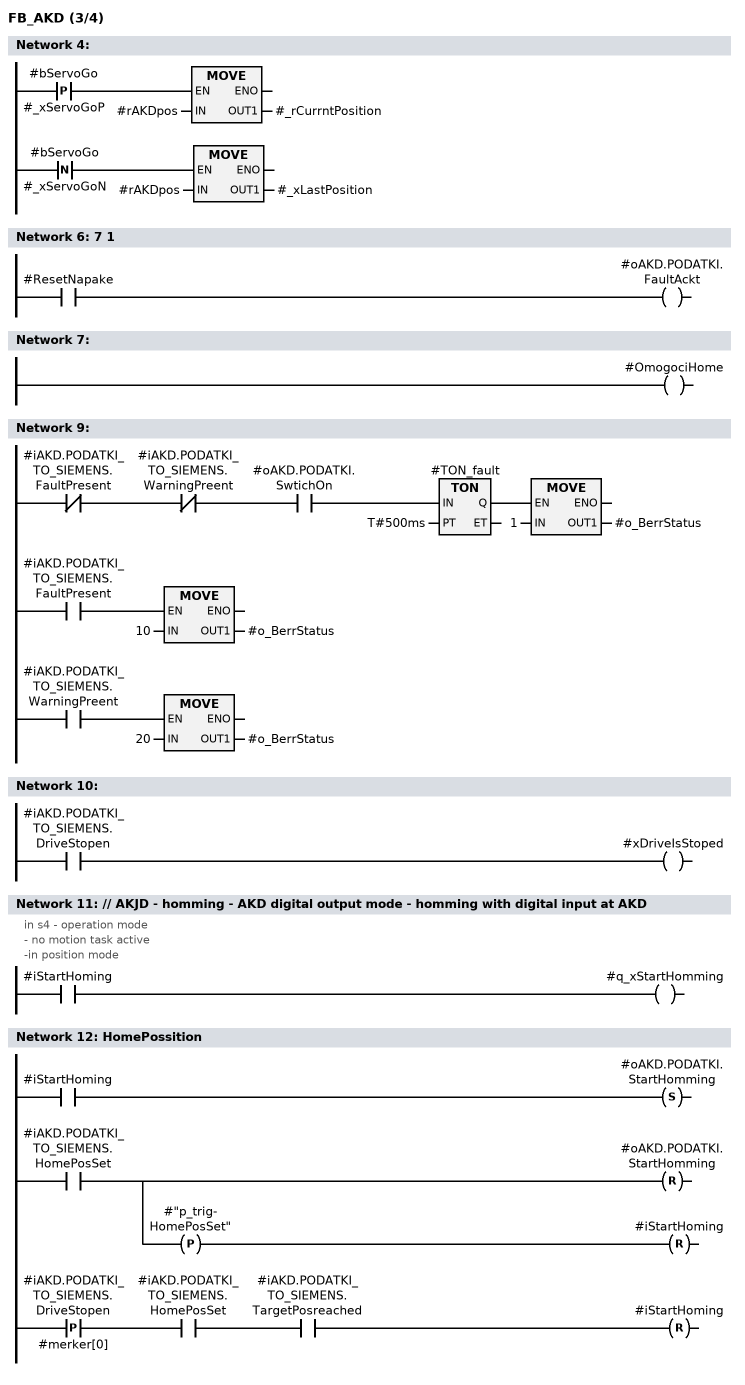
   RUNG wire#powerrail
      P_Contact(operand := #bServoGo, bit := #_xServoGoP)
      Move(in := #rAKDpos, out1 => #_rCurrntPosition)
   END_RUNG
   RUNG wire#powerrail
      N_Contact(operand := #bServoGo, bit := #_xServoGoN)
      Move(in := #rAKDpos, out1 => #_xLastPosition)
   END_RUNG
   // the same network as SCL:
   #_w1 := #bServoGo AND NOT #_xServoGoP;   // rising edge of #bServoGo
   #_xServoGoP := #bServoGo;
   IF #_w1 THEN #_rCurrntPosition := #rAKDpos; END_IF;
   #_w2 := NOT #bServoGo AND #_xServoGoN;   // falling edge of #bServoGo
   #_xServoGoN := #bServoGo;
   IF #_w2 THEN #_xLastPosition := #rAKDpos; END_IF;
END_REGION

REGION Network 5 (SCL)
   //PretvorbaHitrosti
   #diHitrost := INT_TO_REAL(#iNastavitevHitrosti);
   #dwHitrostRez :=((#diHitrost * 4294967295/12000));
   #oAKD.PODATKI.MDI_VELOCITY := REAL_TO_DINT(#dwHitrostRez); //hitrost


   // Operation mode
   #oAKD.PODATKI.MDI_MOD := 16#00_00; //0 - relativni 1//aboslutni gib
   #oAKD.PODATKI.SATANW := #iStPrograma;   //OutputTask

   //pretvorba poziij
   #AKDcurrPos := (#iAKD.PODATKI_TO_SIEMENS.ActualPos * 5 )/ 65536;
   #rAKDpos:= (#iAKD.PODATKI_TO_SIEMENS.ActualPos) / 65536.00;
   //nastavljanjePozicije
   //nastavljanje pozicije
   #oAKD.PODATKI.MDI_TARPOS := (65536 * #dNastavitevPozicije / 5);
END_REGION

REGION Network 6: 7 1
   RUNG wire#powerrail
      Contact( #ResetNapake )
      Coil( #oAKD.PODATKI.FaultAckt )
   END_RUNG
   // the same network as SCL:
   #oAKD.PODATKI.FaultAckt := #ResetNapake;
END_REGION

REGION Network 7
   RUNG wire#powerrail
      Coil( #OmogociHome )
   END_RUNG
   // the same network as SCL:
   #OmogociHome := TRUE;
END_REGION

REGION Network 8: ERROR STATUS
END_REGION

REGION Network 9
   #TON_fault(IN := NOT #iAKD.PODATKI_TO_SIEMENS.FaultPresent AND NOT #iAKD.PODATKI_TO_SIEMENS.WarningPreent AND #oAKD.PODATKI.SwtichOn,   // TON
              PT := T#500ms);
   IF #TON_fault.Q THEN #o_BerrStatus := 1; END_IF;
   IF #iAKD.PODATKI_TO_SIEMENS.FaultPresent THEN #o_BerrStatus := 10; END_IF;
   IF #iAKD.PODATKI_TO_SIEMENS.WarningPreent THEN #o_BerrStatus := 20; END_IF;
END_REGION

REGION Network 10
   RUNG wire#powerrail
      Contact( #iAKD.PODATKI_TO_SIEMENS.DriveStopen )
      Coil( #xDriveIsStoped )
   END_RUNG
   // the same network as SCL:
   #xDriveIsStoped := #iAKD.PODATKI_TO_SIEMENS.DriveStopen;
END_REGION

REGION Network 11: // AKJD - homming - AKD digital output mode - homming with digital input at AKD
   // in s4 - operation mode
   // - no motion task active
   // -in position mode
   RUNG wire#powerrail
      Contact( #iStartHoming )
      Coil( #q_xStartHomming )
   END_RUNG
   // the same network as SCL:
   #q_xStartHomming := #iStartHoming;
END_REGION

REGION Network 12: HomePossition
   RUNG wire#powerrail
      Contact( #iStartHoming )
      S_Coil( #oAKD.PODATKI.StartHomming )
   END_RUNG
   RUNG wire#powerrail
      Contact( #iAKD.PODATKI_TO_SIEMENS.HomePosSet )
      wire#w1
      R_Coil( #oAKD.PODATKI.StartHomming )
   END_RUNG
   RUNG wire#w1
      P_Trig( #"p_trig-HomePosSet" )
      R_Coil( #iStartHoming )
   END_RUNG
   RUNG wire#powerrail
      P_Contact(operand := #iAKD.PODATKI_TO_SIEMENS.DriveStopen, bit := #merker[0])
      Contact( #iAKD.PODATKI_TO_SIEMENS.HomePosSet )
      Contact( #iAKD.PODATKI_TO_SIEMENS.TargetPosreached )
      R_Coil( #iStartHoming )
   END_RUNG
   // the same network as SCL:
   IF #iStartHoming THEN #oAKD.PODATKI.StartHomming := TRUE; END_IF;
   IF #iAKD.PODATKI_TO_SIEMENS.HomePosSet THEN #oAKD.PODATKI.StartHomming := FALSE; END_IF;
   #_w1 := #iAKD.PODATKI_TO_SIEMENS.HomePosSet AND NOT #"p_trig-HomePosSet";   // rising edge
   #"p_trig-HomePosSet" := #iAKD.PODATKI_TO_SIEMENS.HomePosSet;
   IF #_w1 THEN #iStartHoming := FALSE; END_IF;
   #_w2 := #iAKD.PODATKI_TO_SIEMENS.DriveStopen AND NOT #merker[0];   // rising edge of #iAKD.PODATKI_TO_SIEMENS.DriveStopen
   #merker[0] := #iAKD.PODATKI_TO_SIEMENS.DriveStopen;
   IF #_w2 AND #iAKD.PODATKI_TO_SIEMENS.HomePosSet AND #iAKD.PODATKI_TO_SIEMENS.TargetPosreached THEN
       #iStartHoming := FALSE;
   END_IF;
END_REGION

REGION Network 13: OUTPUT : is hommed
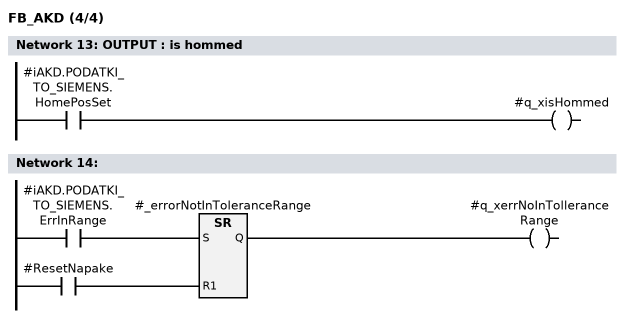
   RUNG wire#powerrail
      Contact( #iAKD.PODATKI_TO_SIEMENS.HomePosSet )
      Coil( #q_xisHommed )
   END_RUNG
   // the same network as SCL:
   #q_xisHommed := #iAKD.PODATKI_TO_SIEMENS.HomePosSet;
END_REGION

REGION Network 14
   RUNG wire#powerrail
      Contact( #iAKD.PODATKI_TO_SIEMENS.ErrInRange )
      S_SR(operand := #_errorNotInToleranceRange, r1 := wire#w1)
      Coil( #q_xerrNoInTolleranceRange )
   END_RUNG
   RUNG wire#powerrail
      Contact( #ResetNapake )
   END_RUNG wire#w1
   // the same network as SCL:
   IF #iAKD.PODATKI_TO_SIEMENS.ErrInRange THEN
       #_errorNotInToleranceRange := TRUE;   // SR flip-flop
   END_IF;
   IF #ResetNapake THEN #_errorNotInToleranceRange := FALSE; END_IF;
   #q_xerrNoInTolleranceRange := #_errorNotInToleranceRange;
END_REGION
END_FUNCTION_BLOCK

FUNCTION_BLOCK "AKD_PN_TG400_v05"   // FB14, SCL
TITLE = AKD_PN_TG400_TIA13_v05
{ S7_Optimized_Access := 'FALSE' }
AUTHOR : jcoleman
FAMILY : TG400
VERSION : 5.0
// This function block supports Profinet communication with the AKD drive using Telegram 400.  It is written in TIA V13. 
// For more information, please see the AKD Profinet Manual and the supporting documentation for this function block.
   VAR_INPUT
      iID : Hw_Io;   // Hardware identifier
      iInit : Bool;   // initialize config for TG400
      iEStop : Bool;   // immediate quick stop and disable
      iSW_Enable : Bool;   // enable/disable
      iStop : Bool;   // stop all movement
      iReset : Bool;   // reset drive faults
      iStart_Homing : Bool;   // start homing
      iStart_Jog : Bool;   // start jog
      iStart_Move : Bool;   // start motion task
      iMT_Pause : Bool;   // pause active motion task
      iMT_MoveType : Word;   // motion task control word 0 = relative; 1 = absolute
      iMTNum : Word;   // motion task number 0x8000 = direct motion task
      iCmdPos : DWord;   // commanded position for motion task or homing
      iCmdVel : DWord;   // commanded velocity for jog or direct motion task
      iCmdAcc : Word;   // commanded acceleration for jog or direct motion task
      iCmdDec : Word;   // commanded deceleration for jog or direct motion task
   END_VAR
   VAR_OUTPUT
      oInitDone : Bool;   // initialization status - 0 while configuring TG400, 1= done
      oStatus : DWord;   // ZSW1
      oPos : DWord;   // actual position
      oVel : Word;   // actual velocity x * 12000 rpm / 2^15
      oCurrent : Word;   // actual current x *DRV.IPEAK / 2^14
      oEnabled : Bool;   // Drive power on
      oError : Bool;   // fault in function block or communication
      oMoving : Bool;   // axis enabled and moving
      oHomed : Bool;   // axis homed
      oInPos : Bool;   // axis within in-position window
      oFault : Bool;   // drive fault
      oWarning : Bool;   // drive warning
   END_VAR
   VAR
      TG_400 : "UDT_AKD_TG400";
      wPNReadStatus : Word;
      bPNReadError : Bool;
      wPNWriteStatus : Word;
      bPNWriteError : Bool;
      bResetDone : Bool;
      bHomeStarted : Bool;
      bStartMoveDone : Bool;
      bEstop : Bool;
      wStartReset : Int;
      wStartMove : Int;
      wSDOStatus : Word;
      bySDODataArray : Array[0..63] of Byte;
      SDOWrite : WRREC;
      SDORead : RDREC;
      bSDOReq : Bool;
      bSDOWriteBusy : Bool;
      bSDOWriteDone : Bool;
      bSDOWriteError : Bool;
      bSDOReadBusy : Bool;
      bSDOReadDone : Bool;
      bSDOReadError : Bool;
      wSDOReadValue : Word;
      wSDOAddress : Word;
      bSWEnabled : Bool;
      wHomingStartPoint : Word;
      bStartMove : Bool;
      bSDOStatusReadActive : Bool;
   END_VAR
BEGIN
   ////////////////////////////////////////////////////////////////////////////////////////////////////////
   // Standard communication module between a Kollmorgen AKD and S7-1200/1500 PLC
   //
   // Version  When        Who         What
   // ---------------------------------------------
   // V 05     09.05.17    JColeman KM Changed Telegram 400 mapping PNU writes to be individual writes, rather
   //                                  than a block write...to be more robust.
   // V 04     08.31.17    JColeman KM Changed error handling to indicate internal block errors.
   // V 03     06.05.17    JColeman KM Changed EStop code to set flag without waiting for motion to stop. 
   //                                  Added setting opmode=2 in init section.
   //                                  Added comments.
   //                                  Added information to FB properties.
   //                                  Turn on real-time jog mode during enable process.
   //                                  Do not use Optimized block access.
   // V 02     05.12.17    JColeman KM Changed names of inputs and outputs to be more user friendly
   //                                  Added output oInitDone to indicate when the telegram configuration is complete
   //                                  Changed name of FB to be specific to TG400
   //                                  Changed verion numbering
   // V 1.000  17.09.15    MRupf KM    Conversion to TIA V13 SP1
   // V 0.004  09.07.15    MRupf KM    Home_dist changed to DINT variable length
   //          06.07.15    MRupf KM    Fault and Warning read locked angainst interruption
   // V 0.003  05.06.15    MRupf KM    New iStart_MT is only accepted after the ZSW1 Bit 12 is FALSE again
   //          03.06.15    MRupf KM    Handshake to start motion task with ZSW1 Bit 12 and auto reset after 500ms #285
   //          14.04.15    MRupf KM    Init write cases extended to not do endless recall on error
   //                                  Homing start stop bug, #246-250
   //                                  Reset STW1.6/.7 only after two PN cylce #214, 283
   // V 0.002  26.02.15    MRupf KM    Setup Telegramm 400 with HOME.DIST, VL.FB, IL.FB
   //                                  Read Fault and Warning No. if acitve
   //                                  Reset STW if drive fault happens while enabled    
   // V 0.001  18.02.15    MRupf KM    First version
   //////////////////////////////////////////////////////////////////////////////////////////////////////////

   // initialisation
   IF #iInit THEN
       #wSDOStatus := 0;
       #oInitDone := FALSE;    //False during telegram configuration
   END_IF;
   IF #wSDOStatus < 20 THEN //set telegram send data = 0
       #TG_400.Send.STW1 := 0;
       #TG_400.Send.SATZANW := 0;
       #TG_400.Send.STW2 := 0;
       #TG_400.Send.MDI_TARPOS := 0;
       #TG_400.Send.MDI_VELOCITY := 0;
       #TG_400.Send.MDI_ACC := 0;
       #TG_400.Send.MDI_DEC := 0;
       #TG_400.Send.MDI_MOD := 0;

       #bPNReadError := FALSE;
       #bPNWriteError := FALSE;
   END_IF;

   // Do the setup of the Telegram 400
   IF NOT #iInit AND #wSDOStatus < 19 THEN

       // Map Telegram 400 Send
       // Clear the Array and start the request
       IF #wSDOStatus = 0 THEN
           FILL_BLK(IN := 0,
                    COUNT := 64,
                    OUT => #bySDODataArray[0]);
           #bSDOReq := TRUE;
           #bSDOWriteDone := FALSE;
           #wSDOStatus := 1; //proceed to Step 1
       END_IF;
       // setup the array data and start WRREC
       IF #wSDOStatus = 1 THEN //Step 1
           #bySDODataArray[0] := 16#ff; //Request Reference
           #bySDODataArray[1] := 16#02; //2 for write PNU
           #bySDODataArray[2] := 16#00; //Axis# is 0 for AKD
           #bySDODataArray[3] := 16#01; //number of parameters
           // Set PNU 915 subindex 8
           #bySDODataArray[4] := 16#10; //Attribute is 0x10
           #bySDODataArray[5] := 16#01; //Number of elements =1
           #bySDODataArray[6] := 16#03; //0x393 for PNU 915
           #bySDODataArray[7] := 16#93; //PNU 915
           #bySDODataArray[8] := 16#00; //subindex
           #bySDODataArray[9] := 16#08; //subindex 8 for 8th word of telegram
           // To PNU 100 (HOME.DIST)
           #bySDODataArray[10] := 16#42; //Format =0x42 for Word
           #bySDODataArray[11] := 16#01; //Number of values
           #bySDODataArray[12] := 16#00; //data
           #bySDODataArray[13] := 16#64; //data - Signal #100 for HOME.DIST

           #SDOWrite(REQ := #bSDOReq, //do the PNU write
                     ID := #iID,
                     INDEX := 47, //AKD suppors "Record Data 47"
                     LEN := 14,   //data length
                     BUSY => #bSDOWriteBusy,
                     DONE => #bSDOWriteDone,
                     ERROR => #bSDOWriteError,
                     RECORD := #bySDODataArray);
           IF #bSDOWriteBusy THEN
               #bSDOReq := FALSE;
           ELSIF #bSDOWriteDone THEN
               #wSDOStatus := 2; //proceed to Step 2
           END_IF;
       END_IF;

       // Map Telegram 400 Receive
       // Clear the Array and start the request
       IF #wSDOStatus = 2 THEN //Step 2
           FILL_BLK(IN := 0,
                    COUNT := 64,
                    OUT => #bySDODataArray[0]);
           #bSDOReq := TRUE;
           #bSDOWriteDone := FALSE;
           #wSDOStatus := 3; //proceed to Step 3
       END_IF;
       // setup the array data and start WRREC
       IF #wSDOStatus = 3 THEN //Step 3
           #bySDODataArray[0] := 16#fe; //Request Reference
           #bySDODataArray[1] := 16#02; //2 for write PNU
           #bySDODataArray[2] := 16#00; //Axis# is 0 for AKD
           #bySDODataArray[3] := 16#01; // Number of parameters to write at a time
           // Set PNU 916 subindex 0
           #bySDODataArray[4] := 16#10; //Attribute is 0x10
           #bySDODataArray[5] := 16#01; //Number of elements =1
           #bySDODataArray[6] := 16#03; //0x394 for PNU 916
           #bySDODataArray[7] := 16#94; //PNU 916
           #bySDODataArray[8] := 16#00; //subindex
           #bySDODataArray[9] := 16#00; //subindex 0 for 1st word of telegram
           // To PNU 2 (ZSW1)
           #bySDODataArray[10] := 16#42; //Format =0x42 for Word
           #bySDODataArray[11] := 16#01; //Number of values
           #bySDODataArray[12] := 16#00; //data
           #bySDODataArray[13] := 16#02; //data - Signal #2 (0x02) for ZSW1

           #SDOWrite(REQ := #bSDOReq, //do the PNU write
                     ID := #iID,
                     INDEX := 47, //AKD suppors "Record Data 47"
                     LEN := 14,   //data length
                     BUSY => #bSDOWriteBusy,
                     DONE => #bSDOWriteDone,
                     ERROR => #bSDOWriteError,
                     RECORD := #bySDODataArray);
           IF #bSDOWriteBusy THEN
               #bSDOReq := FALSE;
           ELSIF #bSDOWriteDone THEN
               #wSDOStatus := 4; //proceed to Step 4
           END_IF;
       END_IF;

       // Clear the Array and start the request
       IF #wSDOStatus = 4 THEN //Step 4
           FILL_BLK(IN := 0,
                    COUNT := 64,
                    OUT => #bySDODataArray[0]);
           #bSDOReq := TRUE;
           #bSDOWriteDone := FALSE;
           #wSDOStatus := 5; //proceed to Step 5
       END_IF;
       // setup the array data and start WRREC
       IF #wSDOStatus = 5 THEN //Step 5
           #bySDODataArray[0] := 16#fd; //Request Reference
           #bySDODataArray[1] := 16#02; //2 for write PNU
           #bySDODataArray[2] := 16#00; //Axis# is 0 for AKD
           #bySDODataArray[3] := 16#01; // Number of parameters to write at a time
           // Set PNU 916 subindex 1
           #bySDODataArray[4] := 16#10; //Attribute is 0x10
           #bySDODataArray[5] := 16#01; //Number of elements =1
           #bySDODataArray[6] := 16#03; //0x394 for PNU 916
           #bySDODataArray[7] := 16#94; //PNU 916
           #bySDODataArray[8] := 16#00; //subindex
           #bySDODataArray[9] := 16#01; //subindex 1 for 2nd word of telegram
           // To PNU 33 (AKTSATZ)
           #bySDODataArray[10] := 16#42; //Format =0x42 for Word
           #bySDODataArray[11] := 16#01; //Number of values
           #bySDODataArray[12] := 16#00; //data
           #bySDODataArray[13] := 16#21; //data - Signal #33 (0x21) for AKTSATZ

           #SDOWrite(REQ := #bSDOReq, //do the PNU write
                     ID := #iID,
                     INDEX := 47, //AKD suppors "Record Data 47"
                     LEN := 14,   //data length
                     BUSY => #bSDOWriteBusy,
                     DONE => #bSDOWriteDone,
                     ERROR => #bSDOWriteError,
                     RECORD := #bySDODataArray);
           IF #bSDOWriteBusy THEN
               #bSDOReq := FALSE;
           ELSIF #bSDOWriteDone THEN
               #wSDOStatus := 6; //proceed to Step 6
           END_IF;
       END_IF;

       // Clear the Array and start the request
       IF #wSDOStatus = 6 THEN //Step 6
           FILL_BLK(IN := 0,
                    COUNT := 64,
                    OUT => #bySDODataArray[0]);
           #bSDOReq := TRUE;
           #bSDOWriteDone := FALSE;
           #wSDOStatus := 7; //proceed to Step 7
       END_IF;
       // setup the array data and start WRREC
       IF #wSDOStatus = 7 THEN //Step 7
           #bySDODataArray[0] := 16#fc; //Request Reference
           #bySDODataArray[1] := 16#02; //2 for write PNU
           #bySDODataArray[2] := 16#00; //Axis# is 0 for AKD
           #bySDODataArray[3] := 16#01; // Number of parameters to write at a time
           // Set PNU 916 subindex 2
           #bySDODataArray[4] := 16#10; //Attribute is 0x10
           #bySDODataArray[5] := 16#01; //Number of elements =1
           #bySDODataArray[6] := 16#03; //0x394 for PNU 916
           #bySDODataArray[7] := 16#94; //PNU 916
           #bySDODataArray[8] := 16#00; //subindex
           #bySDODataArray[9] := 16#02; //subindex 2 for 3rd word of telegram
           // To PNU 4 (ZSW1)
           #bySDODataArray[10] := 16#42; //Format =0x42 for Word
           #bySDODataArray[11] := 16#01; //Number of values
           #bySDODataArray[12] := 16#00; //data
           #bySDODataArray[13] := 16#04; //data - Signal #4 (0x04) for ZSW2

           #SDOWrite(REQ := #bSDOReq, //do the PNU write
                     ID := #iID,
                     INDEX := 47, //AKD suppors "Record Data 47"
                     LEN := 14,   //data length
                     BUSY => #bSDOWriteBusy,
                     DONE => #bSDOWriteDone,
                     ERROR => #bSDOWriteError,
                     RECORD := #bySDODataArray);
           IF #bSDOWriteBusy THEN
               #bSDOReq := FALSE;
           ELSIF #bSDOWriteDone THEN
               #wSDOStatus := 8; //proceed to Step 8
           END_IF;
       END_IF;

       // Clear the Array and start the request
       IF #wSDOStatus = 8 THEN //Step 8
           FILL_BLK(IN := 0,
                    COUNT := 64,
                    OUT => #bySDODataArray[0]);
           #bSDOReq := TRUE;
           #bSDOWriteDone := FALSE;
           #wSDOStatus := 9; //proceed to Step 9
       END_IF;
       // setup the array data and start WRREC
       IF #wSDOStatus = 9 THEN //Step 9
           #bySDODataArray[0] := 16#fb; //Request Reference
           #bySDODataArray[1] := 16#02; //2 for write PNU
           #bySDODataArray[2] := 16#00; //Axis# is 0 for AKD
           #bySDODataArray[3] := 16#01; // Number of parameters to write at a time
           // Set PNU 916 subindex 3
           #bySDODataArray[4] := 16#10; //Attribute is 0x10
           #bySDODataArray[5] := 16#01; //Number of elements =1
           #bySDODataArray[6] := 16#03; //0x394 for PNU 916
           #bySDODataArray[7] := 16#94; //PNU 916
           #bySDODataArray[8] := 16#00; //subindex
           #bySDODataArray[9] := 16#03; //subindex 3 for 4th word of telegram
           // To PNU 28 (XIST_A)
           #bySDODataArray[10] := 16#42; //Format =0x42 for Word
           #bySDODataArray[11] := 16#01; //Number of values
           #bySDODataArray[12] := 16#00; //data
           #bySDODataArray[13] := 16#1C; //data - Signal #28 (0x1C) for XIST_A

           #SDOWrite(REQ := #bSDOReq, //do the PNU write
                     ID := #iID,
                     INDEX := 47, //AKD suppors "Record Data 47"
                     LEN := 14,   //data length
                     BUSY => #bSDOWriteBusy,
                     DONE => #bSDOWriteDone,
                     ERROR => #bSDOWriteError,
                     RECORD := #bySDODataArray);
           IF #bSDOWriteBusy THEN
               #bSDOReq := FALSE;
           ELSIF #bSDOWriteDone THEN
               #wSDOStatus := 10; //proceed to Step 10
           END_IF;
       END_IF;

       // Clear the Array and start the request
       IF #wSDOStatus = 10 THEN //Step 10
           FILL_BLK(IN := 0,
                    COUNT := 64,
                    OUT => #bySDODataArray[0]);
           #bSDOReq := TRUE;
           #bSDOWriteDone := FALSE;
           #wSDOStatus := 11; //proceed to Step 11
       END_IF;
       // setup the array data and start WRREC
       IF #wSDOStatus = 11 THEN //Step 11
           #bySDODataArray[0] := 16#fa; //Request Reference
           #bySDODataArray[1] := 16#02; //2 for write PNU
           #bySDODataArray[2] := 16#00; //Axis# is 0 for AKD
           #bySDODataArray[3] := 16#01; // Number of parameters to write at a time
           // Set PNU 916 subindex 4
           #bySDODataArray[4] := 16#10; //Attribute is 0x10
           #bySDODataArray[5] := 16#01; //Number of elements =1
           #bySDODataArray[6] := 16#03; //0x394 for PNU 916
           #bySDODataArray[7] := 16#94; //PNU 916
           #bySDODataArray[8] := 16#00; //subindex
           #bySDODataArray[9] := 16#04; //subindex 4 for 5th word of telegram
           // To PNU 6 (NIST_A)
           #bySDODataArray[10] := 16#42; //Format =0x42 for Word
           #bySDODataArray[11] := 16#01; //Number of values
           #bySDODataArray[12] := 16#00; //data
           #bySDODataArray[13] := 16#06; //data - Signal #6 (0x06) for NIST_A (VL.FB)

           #SDOWrite(REQ := #bSDOReq, //do the PNU write
                     ID := #iID,
                     INDEX := 47, //AKD suppors "Record Data 47"
                     LEN := 14,   //data length
                     BUSY => #bSDOWriteBusy,
                     DONE => #bSDOWriteDone,
                     ERROR => #bSDOWriteError,
                     RECORD := #bySDODataArray);
           IF #bSDOWriteBusy THEN
               #bSDOReq := FALSE;
           ELSIF #bSDOWriteDone THEN
               #wSDOStatus := 12; //proceed to Step 12
           END_IF;
       END_IF;

       // Clear the Array and start the request
       IF #wSDOStatus = 12 THEN //Step 12
           FILL_BLK(IN := 0,
                    COUNT := 64,
                    OUT => #bySDODataArray[0]);
           #bSDOReq := TRUE;
           #bSDOWriteDone := FALSE;
           #wSDOStatus := 13; //proceed to Step 13
       END_IF;
       // setup the array data and start WRREC
       IF #wSDOStatus = 13 THEN //Step 13
           #bySDODataArray[0] := 16#f9; //Request Reference
           #bySDODataArray[1] := 16#02; //2 for write PNU
           #bySDODataArray[2] := 16#00; //Axis# is 0 for AKD
           #bySDODataArray[3] := 16#01; // Number of parameters to write at a time
           // Set PNU 916 subindex 5
           #bySDODataArray[4] := 16#10; //Attribute is 0x10
           #bySDODataArray[5] := 16#01; //Number of elements =1
           #bySDODataArray[6] := 16#03; //0x394 for PNU 916
           #bySDODataArray[7] := 16#94; //PNU 916
           #bySDODataArray[8] := 16#00; //subindex
           #bySDODataArray[9] := 16#05; //subindex 5 for 6th word of telegram
           // To PNU 52 (ITIST_GLATT)
           #bySDODataArray[10] := 16#42; //Format =0x42 for Word
           #bySDODataArray[11] := 16#01; //Number of values
           #bySDODataArray[12] := 16#00; //data
           #bySDODataArray[13] := 16#34; //data - Signal #52 (0x34) for ITIST_GLATT (IL.FB)

           #SDOWrite(REQ := #bSDOReq, //do the PNU write
                     ID := #iID,
                     INDEX := 47, //AKD suppors "Record Data 47"
                     LEN := 14,   //data length
                     BUSY => #bSDOWriteBusy,
                     DONE => #bSDOWriteDone,
                     ERROR => #bSDOWriteError,
                     RECORD := #bySDODataArray);
           IF #bSDOWriteBusy THEN
               #bSDOReq := FALSE;
           ELSIF #bSDOWriteDone THEN
               #wSDOStatus := 14; //proceed to Step 14
               //#oInitDone := 1;    //telegram configuration complete
           END_IF;
       END_IF;

       // Set OpMode 
       // Clear the Array and start the request
       IF #wSDOStatus = 14 THEN //Step 14
           FILL_BLK(IN := 0,
                    COUNT := 64,
                    OUT => #bySDODataArray[0]);
           #bSDOReq := TRUE;
           #bSDOWriteDone := FALSE;
           #wSDOStatus := 15; //proceed to Step 15
       END_IF;
       // Set OpMode = 2 Position
       IF #wSDOStatus = 15 THEN //Step 15
           #bySDODataArray[0] := 16#fe; //Request Reference
           #bySDODataArray[1] := 16#02; //2 for write PNU
           #bySDODataArray[2] := 16#00; //Axis# is 0 for AKD
           #bySDODataArray[3] := 16#01; // Number of parameters to write at a time
               // Set PNU 930 subindex 0 (DRV.OPMODE)
           #bySDODataArray[4] := 16#10; //Attribute is 0x10
           #bySDODataArray[5] := 16#01; //Number of elements =1
           #bySDODataArray[6] := 16#03; //0x3A2 for PNU 930 - opmode
           #bySDODataArray[7] := 16#A2; //PNU 930
           #bySDODataArray[8] := 16#00; //subindex 0
           #bySDODataArray[9] := 16#00; //subindex 0
               // To 2 (position mode)
           #bySDODataArray[10] := 16#42; //Format =0x42 for Word
           #bySDODataArray[11] := 16#01; //Number of values
           #bySDODataArray[12] := 16#02; //data
           #bySDODataArray[13] := 16#02; //data - vlaue = 2 for position mode

           #SDOWrite(REQ := #bSDOReq, //do the PNU write
                     ID := #iID,
                     INDEX := 47, //AKD suppors "Record Data 47"
                     LEN := 14,   //data length
                     BUSY => #bSDOWriteBusy,
                     DONE => #bSDOWriteDone,
                     ERROR => #bSDOWriteError,
                     RECORD := #bySDODataArray);
           IF #bSDOWriteBusy THEN
               #bSDOReq := FALSE;
           ELSIF #bSDOWriteDone THEN
               #wSDOStatus := 20; // setup complete - skip to process
               #oInitDone := TRUE;    //telegram configuration complete
           END_IF;
       END_IF;
   END_IF;

   // Read ZSW and set output values
   IF NOT #iInit AND #wSDOStatus > 19 THEN
       #wPNReadStatus := DPRD_DAT(LADDR := #iID,
                                  RECORD => #TG_400.Receive);
       IF #wPNReadStatus = 0 THEN
           #bPNReadError := FALSE;

           #oStatus.%W0 := #TG_400.Receive.ZSW1;
           IF #wSDOStatus > 20 THEN
               #oStatus.%W1 := #wSDOReadValue;
           ELSE
               #oStatus.%W1 := 0;
           END_IF;
           #oPos.%W0 := #TG_400.Receive.XIST_A_1;
           #oPos.%W1 := #TG_400.Receive.XIST_A;
           #oVel := #TG_400.Receive.NIST_A;
           #oCurrent := #TG_400.Receive.ITIST_GLATT;

           #oEnabled := #TG_400.Receive.ZSW1.%X0 AND #TG_400.Receive.ZSW1.%X1 AND #TG_400.Receive.ZSW1.%X2 AND NOT #TG_400.Receive.ZSW1.%X6;
           #oFault := #TG_400.Receive.ZSW1.%X3;
           #oMoving := NOT #TG_400.Receive.ZSW1.%X13 OR #TG_400.Receive.ZSW1.%X14 OR #TG_400.Receive.ZSW1.%X12;
           #oHomed := #TG_400.Receive.ZSW1.%X11;
           IF #TG_400.Send.STW1.%X6 THEN        // Reset the InPos Flag for a minimum of one write cycle
               #oInPos := FALSE;
           ELSE
               #oInPos := #TG_400.Receive.ZSW1.%X10;
           END_IF;
           #oWarning := #TG_400.Receive.ZSW1.%X7;
       ELSE
           #bPNReadError := TRUE;
       END_IF;

   END_IF;

   // Do the write always as the zero Telegramm needs to be send on a init aswell
   #wPNWriteStatus := DPWR_DAT(LADDR := #iID,
                               RECORD := #TG_400.Send);

   // set STW1 and values for the AKD
   IF NOT #iInit AND #wSDOStatus > 19 THEN
       IF #wPNWriteStatus = 0 THEN
           #bPNWriteError := FALSE;

           #TG_400.Send.STW1.%X10 := TRUE;
           IF #TG_400.Receive.ZSW1.%X9 THEN     // PLC has control

               // Do a EStop
               IF #iEStop THEN
                   #TG_400.Send.STW1.%X2 := FALSE;
                   #bEstop := TRUE;
               END_IF;

               // Do a reset
               IF #iReset AND NOT #bResetDone THEN
                   #wSDOStatus := 20;
                   #TG_400.Send.STW1.%X7 := TRUE;
                   #bResetDone := TRUE;
                   #bEstop := FALSE;
                   #wStartReset := #TG_400.Receive.ZSW2;
               END_IF;
               IF ABS(#wStartReset - #TG_400.Receive.ZSW2) > 2 THEN
                   #TG_400.Send.STW1.%X7 := FALSE;
               END_IF;

               // Enable the drive
               IF #iSW_Enable AND NOT #bEstop AND NOT (#bSWEnabled AND #TG_400.Receive.ZSW1.%X6 OR #TG_400.Receive.ZSW1.%X3) THEN
                   IF #TG_400.Receive.ZSW1.%X6 THEN      // Switch on inhibited
                       #TG_400.Send.STW1.%X1 := TRUE;
                       #TG_400.Send.STW1.%X2 := TRUE;
                   ELSE
                       IF #TG_400.Receive.ZSW1.%X0 THEN     // Ready for switiching on
                           #TG_400.Send.STW1.%X0 := TRUE;
                           IF #TG_400.Receive.ZSW1.%X1 THEN       // Switched on
                               #TG_400.Send.STW1.%X3 := TRUE;
                               IF #TG_400.Receive.ZSW1.%X2 THEN       // Operation
                                   #TG_400.Send.STW1.%X12 := TRUE; //turn on real time jogging mode
                                   #bSWEnabled := TRUE;

                                   // Do a Stop
                                   IF #iStop THEN
                                       #TG_400.Send.STW1.%X4 := FALSE;   // Stop active motion task
                                       #TG_400.Send.STW1.%X5 := FALSE;   // Stop active motion task
                                       #TG_400.Send.STW1.%X8 := FALSE;   // Stop jog 1
                                       #TG_400.Send.STW1.%X9 := FALSE;   // Stop jog 2
                                       #TG_400.Send.STW1.%X11 := FALSE;  // Stop homeing
                                       //#TG_400.Send.STW1.%X12 := FALSE;  // Stop real time jogging mode
                                   ELSE

                                       // Do home
                                       IF #iStart_Homing AND NOT #bHomeStarted THEN
                                           #TG_400.Send.HOME_DIST := #iCmdPos.%W1;
                                           #TG_400.Send.HOME_DIST_1 := #iCmdPos.%W0;
                                           #TG_400.Send.STW1.%X11 := TRUE;
                                           #wHomingStartPoint := #TG_400.Receive.ZSW2;
                                           #bHomeStarted := TRUE;
                                       ELSE
                                           IF #TG_400.Receive.ZSW1.%X11 AND #TG_400.Receive.ZSW1.%X13 AND (ABS(#wHomingStartPoint - #TG_400.Receive.ZSW2) > 5) THEN
                                               #TG_400.Send.STW1.%X11 := FALSE;
                                           END_IF;

                                           // Jogging
                                           IF #iStart_Jog AND #iCmdVel <> 0 THEN
                                               #TG_400.Send.STW1.%X8 := TRUE;
                                               //#TG_400.Send.STW1.%X12 := TRUE;

                                               // if the speed input is negative set Bit 13 for reverse direction 
                                               IF #iCmdVel.%X31 = 1 THEN
                                                   #TG_400.Send.STW1.%X13 := TRUE;
                                                   #TG_400.Send.MDI_VELOCITY := (16#ffff - #iCmdVel.%W1 + 1);
                                                   #TG_400.Send.MDI_VELOCITY_1 := (16#ffff - #iCmdVel.%W0 + 1);
                                               ELSE
                                                   #TG_400.Send.STW1.%X13 := FALSE;
                                                   #TG_400.Send.MDI_VELOCITY := #iCmdVel.%W1;
                                                   #TG_400.Send.MDI_VELOCITY_1 := #iCmdVel.%W0;
                                               END_IF;

                                               #TG_400.Send.MDI_ACC := #iCmdAcc;
                                               #TG_400.Send.MDI_DEC := #iCmdDec;
                                           ELSE
                                               #TG_400.Send.STW1.%X8 := FALSE;
                                               //#TG_400.Send.STW1.%X12 := FALSE;

                                               // Interrupt a move
                                               IF #iMT_Pause THEN
                                                   #TG_400.Send.STW1.%X5 := FALSE;    // intermediate stop, motion is paused and will continue when the pause is lifted
                                               ELSE
                                                   #TG_400.Send.STW1.%X5 := TRUE;    // No intermediate stop
                                               END_IF;

                                               // Reset the rising edge of the start bit to be read for the next task
                                               IF #TG_400.Receive.ZSW1.%X12 OR ABS(#wStartMove - #TG_400.Receive.ZSW2) > 62 THEN //if start command has been acknowledged, or >62 telegram transmissions
                                                   #bStartMoveDone := TRUE; // the process to start the move has been completed
                                                   #TG_400.Send.STW1.%X6 := FALSE; //turn off the start bit
                                               END_IF;
                                               // Move
                                               IF #iStart_Move AND NOT #bStartMove THEN
                                                   #TG_400.Send.MDI_MOD := #iMT_MoveType;   // 1 = absolute, 0 = relative
                                                   #TG_400.Send.SATZANW := #iMTNum;      // 0x8000 = direct motion task, otherwise select a motion task from the AKD
                                                   #TG_400.Send.MDI_TARPOS := #iCmdPos.%W1;
                                                   #TG_400.Send.MDI_TARPOS_1 := #iCmdPos.%W0;
                                                   #TG_400.Send.MDI_VELOCITY := #iCmdVel.%W1;
                                                   #TG_400.Send.MDI_VELOCITY_1 := #iCmdVel.%W0;
                                                   #TG_400.Send.MDI_ACC := #iCmdAcc;
                                                   #TG_400.Send.MDI_DEC := #iCmdDec;
                                                   #TG_400.Send.STW1.%X4 := TRUE;    // Do not reject traversing task
                                                   #TG_400.Send.STW1.%X5 := TRUE;    // No intermediate stop
                                                   #TG_400.Send.STW1.%X6 := TRUE;    // Start the move

                                                   #bStartMove := TRUE; // the process to start the move has been started but not completed
                                                   #bStartMoveDone := FALSE; // the process to start the move has not been completed
                                                   #wStartMove := #TG_400.Receive.ZSW2;
                                               END_IF; //If Start move

                                           END_IF; //If Start Jog
                                       END_IF; //If Start Homing
                                   END_IF; // If Stop
                               END_IF; // If ZSW1 bit2 Operation Enabled
                           END_IF; // If ZSW1 bit1 Switched On
                       END_IF; // If ZSW1 bit0 Ready for Switch On
                   END_IF; // If ZSW1 bit6 Switch-On Inhibited

                   // If the axis gets disabled all the corresponding motion signals have to be reset    
               ELSE
                   #bSWEnabled := FALSE;

                   #TG_400.Send.STW1.%X0 := FALSE;
                   #TG_400.Send.STW1.%X1 := FALSE;
                   #TG_400.Send.STW1.%X2 := FALSE;
                   #TG_400.Send.STW1.%X3 := FALSE;
                   #TG_400.Send.STW1.%X4 := FALSE;
                   #TG_400.Send.STW1.%X5 := FALSE;
                   #TG_400.Send.STW1.%X6 := FALSE;
                   #TG_400.Send.STW1.%X8 := FALSE;
                   #TG_400.Send.STW1.%X9 := FALSE;
                   #TG_400.Send.STW1.%X11 := FALSE;
                   #TG_400.Send.STW1.%X12 := FALSE;
               END_IF; //If Enable
           END_IF; // ZSW1 bit9 PLC has control
       ELSE
           #bPNWriteError := TRUE;
       END_IF; //If #wPNWriteStatus = 0

       // Read drive faults and warning on occurens
       IF #oFault THEN
           // If alarm is not read yet: start read
           IF NOT #wSDOStatus.%X6 AND NOT #bSDOStatusReadActive THEN
               #wSDOStatus := 64;
               #wSDOAddress := 16#09AD;     // Read PNU 2477 (DRV.FAULT1)
               #bSDOStatusReadActive := TRUE;
           END_IF;

           // If warning is not read yet: start read
       ELSIF #oWarning THEN
           IF NOT #wSDOStatus.%X5 AND NOT #bSDOStatusReadActive THEN
               #wSDOStatus := 32;
               #wSDOAddress := 16#0AE7;    // Read PNU2791 (DRV.WARNING1)
               #bSDOStatusReadActive := TRUE;
           END_IF;
       ELSE
           IF NOT #bSDOStatusReadActive THEN
               #wSDOStatus := 20;
           END_IF;
       END_IF; //IF #oFault

       // start the reading signal
       IF #wSDOStatus >= 32 THEN
           // Always clean out old values first
           IF #bSDOWriteBusy THEN
               #bSDOReq := FALSE;
           ELSE
               FILL_BLK(IN := 0,
                        COUNT := 64,
                        OUT => #bySDODataArray[0]);
               #bSDOReq := TRUE;
               #bSDOWriteDone := FALSE;
           END_IF;
           // Start the read cylce to the corrsponding PNU 
           IF #wSDOStatus = 32 OR #wSDOStatus = 64 THEN
               #bySDODataArray[0] := #wSDOStatus.%B0;
               #bySDODataArray[1] := 16#01;
               #bySDODataArray[2] := 16#00;
               #bySDODataArray[3] := 16#01;

               #bySDODataArray[4] := 16#10;
               #bySDODataArray[5] := 16#01;
               #bySDODataArray[6] := #wSDOAddress.%B1;
               #bySDODataArray[7] := #wSDOAddress.%B0;
               #bySDODataArray[8] := 16#00;
               #bySDODataArray[9] := 16#00;

               #SDOWrite(REQ := #bSDOReq,
                         ID := #iID,
                         INDEX := 47,
                         LEN := 14,
                         BUSY => #bSDOWriteBusy,
                         DONE => #bSDOWriteDone,
                         ERROR => #bSDOWriteError,
                         RECORD := #bySDODataArray);
               IF #bSDOWriteDone THEN
                   #wSDOStatus := #wSDOStatus + 1;
               END_IF;
           END_IF; //IF #wSDOStatus = 32 OR #wSDOStatus = 64

           // read the value back
           IF #wSDOStatus = 33 OR #wSDOStatus = 65 THEN
               #SDORead(REQ := #bSDOReq,
                        ID := #iID,
                        INDEX := 47,
                        MLEN := 14,
                        BUSY => #bSDOReadBusy,
                        VALID => #bSDOReadDone,
                        ERROR => #bSDOReadError,
                        RECORD := #bySDODataArray);
               IF #bSDOReadDone THEN
                   IF #bySDODataArray[4] = 66 THEN               // if the read signal is a Word use Byte 6&7
                       #wSDOReadValue.%B0 := #bySDODataArray[7];
                       #wSDOReadValue.%B1 := #bySDODataArray[6];
                   ELSE                                        // if the read signal is a DWord use Byte 8&9
                       #wSDOReadValue.%B0 := #bySDODataArray[9];
                       #wSDOReadValue.%B1 := #bySDODataArray[8];
                   END_IF;
                   IF #wSDOReadValue = 0 THEN  // If the read value is zero repeat the read cycle
                       #wSDOStatus := #wSDOStatus - 1;
                   ELSE
                       #wSDOStatus := #wSDOStatus + 1;
                       #bSDOStatusReadActive := FALSE;
                   END_IF;
               END_IF; //IF #bSDOReadDone
           END_IF; //IF #wSDOStatus = 33 OR #wSDOStatus = 65
       END_IF; //IF #wSDOStatus >= 32
   END_IF; //IF NOT #iInit AND #wSDOStatus > 19

   //  check for rising edge for the input parameters
   IF NOT #iReset AND #bResetDone THEN
       #bResetDone := FALSE;
   END_IF;
   IF NOT #iStart_Homing AND #bHomeStarted THEN
       #bHomeStarted := FALSE;
   END_IF;
   IF NOT #iStart_Move AND #bStartMove AND #bStartMoveDone AND NOT #TG_400.Receive.ZSW1.%X12 THEN
       #bStartMove := FALSE;
       #bStartMoveDone := FALSE;
   END_IF;

   // fault detection/handling within the bloc
   IF #bPNReadError OR #bPNWriteError OR #bSDOReadError OR #bSDOWriteError THEN
       #oError := TRUE;
       IF #bPNReadError THEN
           #oStatus := #wPNReadStatus; //indicates internal FB error
       END_IF;
       IF #bPNWriteError THEN
           #oStatus := #wPNWriteStatus; //indicates internal FB error
       END_IF;
   ELSIF #wSDOStatus > 19 THEN
       #oError := FALSE;
   END_IF;
END_FUNCTION_BLOCK

// folder: AKD/PNU

